REGION Network 3: Falha de comando
   RUNG wire#powerrail
      Contact( #TEMP0 )
      wire#w1
      S_Coil( #YFPP )
   END_RUNG
   RUNG wire#powerrail
      Contact( #TEMP1 )
   END_RUNG wire#w1
   RUNG wire#w1
      Coil( #AUX01 )
   END_RUNG
   // the same network as SCL:
   #_w1 := #TEMP0 OR #TEMP1;
   IF #_w1 THEN #YFPP := TRUE; END_IF;
   #AUX01 := #_w1;
END_REGION

REGION Network 4: Reset falha no acionamento
   RUNG wire#powerrail
      Contact( #CRF )
      I_Contact( #AUX01 )
      wire#w1
      R_Coil( #YFPP )
   END_RUNG
   RUNG wire#powerrail
      I_Contact( #DL )
   END_RUNG wire#w1
   // the same network as SCL:
   IF (#CRF AND NOT #AUX01) OR NOT #DL THEN #YFPP := FALSE; END_IF;
END_REGION

REGION Network 5: Falha
   RUNG wire#powerrail
      Contact( #DL )
      Contact( #MF1 )
      Contact( #MF2 )
      I_Contact( #YFPP )
      Not()
      Coil( #YF )
   END_RUNG
   // the same network as SCL:
   #YF := NOT (#DL AND #MF1 AND #MF2 AND NOT #YFPP);
END_REGION

REGION Network 6: Transição automático/manual
   RUNG wire#powerrail
      I_Contact( #CMA )
      P_Trig( #AUX02 )
      Contact( #MR )
      Contact( #ML )
      Coil( #AUX03 )
   END_RUNG
   // the same network as SCL:
   #_w1 := NOT #CMA AND NOT #AUX02;   // rising edge
   #AUX02 := NOT #CMA;
   #AUX03 := #_w1 AND #MR AND #ML;
END_REGION

REGION Network 7: Liga em manual
   RUNG wire#powerrail
      Contact( #CLM )
      wire#w1
      I_Contact( #CMA )
      I_Contact( #CDM )
      I_Contact( #YF )
      Contact( #HM )
      Contact( #MR )
      Coil( #AUX04 )
   END_RUNG
   RUNG wire#powerrail
      Contact( #AUX04 )
   END_RUNG wire#w1
   RUNG wire#powerrail
      Contact( #AUX03 )
   END_RUNG wire#w1
   // the same network as SCL:
   #AUX04 := (#CLM OR #AUX04 OR #AUX03) AND NOT #CMA AND NOT #CDM AND NOT #YF AND #HM AND #MR;
END_REGION

REGION Network 8: Liga em automático
   RUNG wire#powerrail
      Contact( #CMA )
      I_Contact( #YF )
      Contact( #HA )
      Contact( #MR )
      Coil( #AUX05 )
   END_RUNG
   // the same network as SCL:
   #AUX05 := #CMA AND NOT #YF AND #HA AND #MR;
END_REGION

REGION Network 9: Comando liga motor
   RUNG wire#powerrail
      Contact( #AUX05 )
      wire#w1
      Coil( #CL )
   END_RUNG
   RUNG wire#powerrail
      Contact( #AUX04 )
   END_RUNG wire#w1
   // the same network as SCL:
   #CL := #AUX05 OR #AUX04;
END_REGION

REGION Network 10
   RUNG wire#powerrail
      Contact( "AlwaysTRUE" )
      wire#w1
      Contact( #CL1S )
      Contact( #ML )
      P_Trig( #AUX06 )
      { S7_Templates := "SrcType := Int"; S7_GenerateENO := "TRUE" } Add(in1 := #SEG, in2 := 1, out => #SEG)
   END_RUNG
   RUNG wire#w1
      { S7_Templates := "SrcType := Int" } GE_Contact(in1 := #SEG, in2 := 60)
      P_Trig( #P60S )
      Coil( #AUX07 )
   END_RUNG
   // the same network as SCL:
   #_w1 := "AlwaysTRUE" AND #CL1S AND #ML;
   #_w2 := #_w1 AND NOT #AUX06;   // rising edge
   #AUX06 := #_w1;
   IF #_w2 THEN #SEG := #SEG + 1; END_IF;
   #_w3 := "AlwaysTRUE" AND (#SEG >= 60);
   #_w4 := #_w3 AND NOT #P60S;   // rising edge
   #P60S := #_w3;
   #AUX07 := #_w4;
END_REGION

REGION Network 11
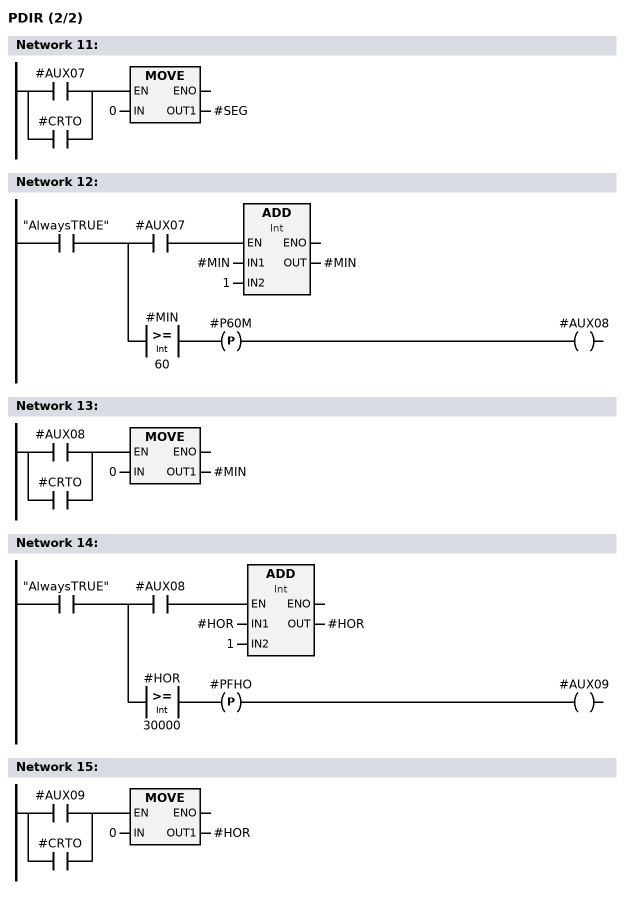
   RUNG wire#powerrail
      Contact( #AUX07 )
      wire#w1
      { S7_GenerateENO := "TRUE" } Move(in := 0, out1 => #SEG)
   END_RUNG
   RUNG wire#powerrail
      Contact( #CRTO )
   END_RUNG wire#w1
   // the same network as SCL:
   IF #AUX07 OR #CRTO THEN #SEG := 0; END_IF;
END_REGION

REGION Network 12
   RUNG wire#powerrail
      Contact( "AlwaysTRUE" )
      wire#w1
      Contact( #AUX07 )
      { S7_Templates := "SrcType := Int"; S7_GenerateENO := "TRUE" } Add(in1 := #MIN, in2 := 1, out => #MIN)
   END_RUNG
   RUNG wire#w1
      { S7_Templates := "SrcType := Int" } GE_Contact(in1 := #MIN, in2 := 60)
      P_Trig( #P60M )
      Coil( #AUX08 )
   END_RUNG
   // the same network as SCL:
   IF "AlwaysTRUE" AND #AUX07 THEN #MIN := #MIN + 1; END_IF;
   #_w1 := "AlwaysTRUE" AND (#MIN >= 60);
   #_w2 := #_w1 AND NOT #P60M;   // rising edge
   #P60M := #_w1;
   #AUX08 := #_w2;
END_REGION

REGION Network 13
   RUNG wire#powerrail
      Contact( #AUX08 )
      wire#w1
      { S7_GenerateENO := "TRUE" } Move(in := 0, out1 => #MIN)
   END_RUNG
   RUNG wire#powerrail
      Contact( #CRTO )
   END_RUNG wire#w1
   // the same network as SCL:
   IF #AUX08 OR #CRTO THEN #MIN := 0; END_IF;
END_REGION

REGION Network 14
   RUNG wire#powerrail
      Contact( "AlwaysTRUE" )
      wire#w1
      Contact( #AUX08 )
      { S7_Templates := "SrcType := Int"; S7_GenerateENO := "TRUE" } Add(in1 := #HOR, in2 := 1, out => #HOR)
   END_RUNG
   RUNG wire#w1
      { S7_Templates := "SrcType := Int" } GE_Contact(in1 := #HOR, in2 := 30000)
      P_Trig( #PFHO )
      Coil( #AUX09 )
   END_RUNG
   // the same network as SCL:
   IF "AlwaysTRUE" AND #AUX08 THEN #HOR := #HOR + 1; END_IF;
   #_w1 := "AlwaysTRUE" AND (#HOR >= 30000);
   #_w2 := #_w1 AND NOT #PFHO;   // rising edge
   #PFHO := #_w1;
   #AUX09 := #_w2;
END_REGION

REGION Network 15
   RUNG wire#powerrail
      Contact( #AUX09 )
      wire#w1
      { S7_GenerateENO := "TRUE" } Move(in := 0, out1 => #HOR)
   END_RUNG
   RUNG wire#powerrail
      Contact( #CRTO )
   END_RUNG wire#w1
   // the same network as SCL:
   IF #AUX09 OR #CRTO THEN #HOR := 0; END_IF;
END_REGION
END_FUNCTION_BLOCK

FUNCTION "ALARME" : Void   // FC2, SCL
{ S7_Optimized_Access := 'TRUE' }
VERSION : 0.1
BEGIN
   REGION "ALARMES IHM"
       // Statement section REGION
       "ALM0" := %DB300.DBW0;
       "ALM2" := %DB300.DBW2;
       "ALM4" := %DB300.DBW4;
       "ALM6" := %DB300.DBW6;
       "ALM8" := %DB300.DBW8;
       "ALM10" := %DB300.DBW10;
       "ALM12" := %DB300.DBW12;
       "ALM14" := %DB300.DBW14;
       "ALM16" := %DB300.DBW16;
   END_REGION
END_FUNCTION

FUNCTION "IO" : Void   // FC4, SCL
{ S7_Optimized_Access := 'TRUE' }
VERSION : 0.1
BEGIN
   REGION "Status e alarme elevatória principal 1"
       // Statement section REGION
       "Digitais"."MB-01-YFI" := "MB_01_DINV";
       "Digitais"."MB-01-YFB" := "MB_01_DMB";
       "Digitais"."MB-01-YFF" :="MB_01_FF";
       "Digitais"."MB-01-EMER" := NOT "MB_01_EMER";
       "Digitais"."MB-01-ML" :="MB_01_ML";
       "Digitais"."MB-01-YSH" :="MB_01_BL" OR "MB_01_SH";
       "Digitais"."MB-01-MM" :="MB_01_MMNT";
       "Digitais"."MB-01-MA" :="MB_01_MA";
       "Digitais"."MB-01-MN" :="MB_01_MN";
       "Digitais"."MB-01-HM" :="MB_01_HMNT";
       "Digitais"."MB-01-RST" :="MB_01_RST";
       "Digitais"."MB-01-INTRU" :="MB_01_INTRU";

       "MB_01_RR" :="COMANDOS"."MB-01-HS4";
       "MB_01_INTV" :="DIVERSOS"."MB-01-SP";
       "MB_01_INTVS" :="DIVERSOS"."MB-01-SP";


   END_REGION
   REGION "Status e alarme elevatória principal 2"
       // Statement section REGION
       "Digitais"."MB-02-YFI" := "MB_02_DINV";
       "Digitais"."MB-02-YFB" := "MB_02_DMB";
       "Digitais"."MB-02-YFF" := "MB_02_FF";
       "Digitais"."MB-02-EMER" := NOT "MB_02_EMER";
       "Digitais"."MB-02-ML" := "MB_02_ML";
       "Digitais"."MB-02-YSH" := "MB_02_BL" OR "MB_02_SH";
       "Digitais"."MB-02-MM" := "MB_02_MMNT";
       "Digitais"."MB-02-MA" := "MB_02_MA";
       "Digitais"."MB-02-MN" := "MB_02_MN";
       "Digitais"."MB-02-HM" := "MB_02_HMNT";
       "Digitais"."MB-02-RST" := "MB_02_RST";
       "Digitais"."MB-02-INTRU" := "MB_02_INTRU";

       "MB_02_RR" := "COMANDOS"."MB-02-HS4";
       "MB_02_INTV" := "DIVERSOS"."MB-02-SP";
       "MB_02_INTVS" := "DIVERSOS"."MB-02-SP";


   END_REGION
   REGION "Status e alarme elevatória principal 3"
       // Statement section REGION
       "Digitais"."MB-03-YFI" := "MB_03_DINV";
       "Digitais"."MB-03-YFB" := "MB_03_DMB";
       "Digitais"."MB-03-YFF" := "MB_03_FF";
       "Digitais"."MB-03-EMER" := NOT "MB_03_EMER";
       "Digitais"."MB-03-ML" := "MB_03_ML";
       "Digitais"."MB-03-YSH" := "MB_03_BL" OR "MB_03_SH";
       "Digitais"."MB-03-MM" := "MB_03_MMNT";
       "Digitais"."MB-03-MA" := "MB_03_MA";
       "Digitais"."MB-03-MN" := "MB_03_MN";
       "Digitais"."MB-03-HM" := "MB_03_HMNT";
       "Digitais"."MB-03-RST" := "MB_03_RST";
       "Digitais"."MB-03-INTRU" := "MB_03_INTRU";

       "MB_03_RR" := "COMANDOS"."MB-03-HS4";
       "MB_03_INTV" := "DIVERSOS"."MB-03-SP";
       "MB_03_INTVS" := "DIVERSOS"."MB-03-SP";


   END_REGION
   REGION "Status e alarme elevatória principal 4"
       // Statement section REGION
       "Digitais"."MB-04-YFI" := "MB_04_DINV";
       "Digitais"."MB-04-YFB" := "MB_04_DMB";
       "Digitais"."MB-04-YFF" := "MB_04_FF";
       "Digitais"."MB-04-EMER" := NOT "MB_04_EMER";
       "Digitais"."MB-04-ML" := "MB_04_ML";
       "Digitais"."MB-04-YSH" := "MB_04_BL" OR "MB_04_SH";
       "Digitais"."MB-04-MM" := "MB_04_MMNT";
       "Digitais"."MB-04-MA" := "MB_04_MA";
       "Digitais"."MB-04-MN" := "MB_04_MN";
       "Digitais"."MB-04-HM" := "MB_04_HMNT";
       "Digitais"."MB-04-RST" := "MB_04_RST";
       "Digitais"."MB-04-INTRU" := "MB_04_INTRU";

       "MB_04_RR" := "COMANDOS"."MB-04-HS4";
       "MB_04_INTV" := "DIVERSOS"."MB-04-SP";
       "MB_04_INTVS" := "DIVERSOS"."MB-04-SP";


   END_REGION

   REGION "Status e alarme PCM-E-CF-01-04"
       // Statement section REGION
       "Digitais".PCM_EEE_EMER := NOT "PCM_EEE_EMER";
       "Digitais".PCM_EEE_K27 := "PCM_EEE_K27";
       "Digitais".PCM_EEE_DISJ_LIG := "PCM_EEE_DJL";
       "Digitais".PCM_EEE_DISJ_DESLIG := "PCM_EEE_DJD";
       "Digitais".PCM_EEE_DISJ_YFAL := "PCM_EEE_DJYFAL";
       "Digitais".PCM_EEE_DISJ_FAL_GR := "PCM_EEE_DJFG";
       "Digitais".PCM_EEE_TR01_KA3 := "PCM_EEE_TR01_KA3";
       "Digitais".PCM_EEE_TR01_KA4 := "PCM_EEE_TR01_KA4";
       "Digitais".PCM_EEE_TR01_KA5 := "PCM_EEE_TR01_KA5";
       "Digitais".PCM_EEE_INTRU := "PCM_EEE_INTRU";
   END_REGION

   REGION "Status e alarme QGBT-AUX-01"
       // Statement section REGION
       "Digitais".QGBT_EMER := NOT "QGBT_EMER";
       "Digitais".QGBT_K27 := "QGBT_K27";
       "Digitais".QGBT_DJL := "QGBT_DISJ_LIG";
       "Digitais".QGBT_DJD := "QGBT_DISJ_DESLIG";
       "Digitais".QGBT_DJYFAL := "QGBT_DISJ_YFAL";
       "Digitais".QGBT_INTRU := "QGBT_INTRU";
   END_REGION

   REGION "CHAVE DE NIVEL LS-001"
       // Statement section REGION
       // 
       "DIVERSOS".TMR[5].TON(IN := "LSL_001",
                             PT := T#5S);
       "DIVERSOS".TMR[6].TON(IN := "LSH_001",
                             PT := T#5S);
       "Digitais".LSL_001 := "DIVERSOS".TMR[5].Q;
       "Digitais".LSH_001 := "DIVERSOS".TMR[6].Q;
   END_REGION

   REGION "CHAVE DE NIVEL LS-002"
       // Statement section REGION
       "DIVERSOS".TMR[7].TON(IN := "LSL_002",
                             PT := T#5S);
       "DIVERSOS".TMR[8].TON(IN := "LSH_002",
                             PT := T#5S);
       "Digitais".LSL_002 := "DIVERSOS".TMR[7].Q;
       "Digitais".LSH_002 := "DIVERSOS".TMR[8].Q;
   END_REGION

   REGION "Status e alarme PCE-EEE"
       // Statement section REGION
       "Digitais".PCE_EEE_INTRU := "PCE_EEE_INTRU";
       "Digitais".PCE_EEE_UPS_ALM := "PCE_EEE_UPS_ALM";
       "Digitais".PCE_EEE_UPS_FE := "PCE_EEE_UPS_FE";
       "Digitais".PCE_EEE_UPS_CHAR := "PCE_EEE_UPS_CHAR";






   END_REGION
END_FUNCTION

FUNCTION "MB-01" : Void   // FC7, SCL
{ S7_Optimized_Access := 'TRUE' }
VERSION : 0.1
   VAR_TEMP
      IM : Bool;   // Intertravamento manual = 0
      IA : Bool;   // Intertravamento automáticol = 0
      HABM : Bool;   // Habilita funcionamento manual = 1
      HABA : Bool;   // Habilita funcionamento automático = 1
      CLM : Bool;   // Comando liga motor
      PROT : Bool;   // Proteção do motor acionada
   END_VAR
BEGIN
   REGION Intertravamento maual/automático
       // Statement section REGION
       IF (NOT "Digitais".QGBT_EMER AND NOT "Digitais".PCM_EEE_EMER AND NOT "Digitais"."MB-01-EMER") = 1 THEN
           // Statement section IF
           #IA := 1;
           #IM := 1;
       ELSE
           #IA := 0;
           #IM := 0;
       END_IF;

   END_REGION

   REGION Habilita funcionamento automático
       // Statement section REGION
       IF (#IA AND "DIVERSOS"."MB-01-SP") = 1 THEN
           // Statement section IF
           #HABA := 1;
       ELSE
           #HABA := 0;
       END_IF;

   END_REGION

   REGION Habilita funcionamento manual
       // Statement section REGION
       IF #IM THEN
           // Statement section IF
           #HABM := 1;
       ELSE
           #HABM := 0;
       END_IF;
   END_REGION

   REGION Bloco de acionamento DO motor
       // Statement section REGION
       "PDIR_DB_MB-01"(ML:="Digitais"."MB-01-YSH",
                       MR:="Digitais"."MB-01-YR",
                       DL:=NOT "Digitais"."MB-01-YFI" AND NOT "Digitais"."MB-01-YFB" AND NOT "Digitais"."MB-01-YFF",
                       MF1:="AlwaysTRUE",
                       MF2:="AlwaysTRUE",
                       HM:=#HABM,
                       HA:=#HABA,
                       CMA:="COMANDOS"."MB-01-HS1",
                       CLM:="COMANDOS"."MB-01-HS2",
                       CDM:="COMANDOS"."MB-01-HS3",
                       CRF:="COMANDOS"."MB-01-HS4" OR "Digitais"."MB-01-RST",
                       CRTO:="COMANDOS"."MB-01-HS5",
                       CL1S:="Clock_1Hz",
                       YFPP=>"Digitais"."MB-01-YFA",
                       YF=>"Digitais"."MB-01-YF",
                       CL=>"MB_01_SH",
                       SEG:="Totalizadores"."MB-01-SO",
                       MIN:="Totalizadores"."MB-01-MO",
                       HOR:="Totalizadores"."MB-01-HO");

                    END_REGION

   REGION Reset dos comandos de pulso
       // Statement section REGION
       IF "COMANDOS"."MB-01-HS2" THEN
           // Statement section IF
           "COMANDOS"."MB-01-HS2" := 0;
       END_IF;
       IF "COMANDOS"."MB-01-HS3" THEN
           // Statement section IF
           "COMANDOS"."MB-01-HS3" := 0;
       END_IF;
       IF "COMANDOS"."MB-01-HS4" THEN
           // Statement section IF
           "COMANDOS"."MB-01-HS4" := 0;
       END_IF;
       IF "COMANDOS"."MB-01-HS5" THEN
           // Statement section IF
           "COMANDOS"."MB-01-HS5" := 0;
       END_IF;
   END_REGION

   REGION Elevatoria principal modo automatico
       IF ("Digitais"."MB-01-MA") = 1 THEN
           "Digitais"."MB-01-YR" := 1;
       ELSE
           "Digitais"."MB-01-YR" := 0;
       END_IF;

   END_REGION

   REGION Proteção hidraulica MB-01
       // Statement section REGION
       IF ("VARIAVEIS".LIT_001 <= "SETPOINTS".SP_NVL_MIN) OR "Digitais".LSL_002 OR "Digitais"."LIT_001-YLL" THEN
           // Statement section IF
           "MB_01_PH" := 1;
       ELSE
           "MB_01_PH" := 0;
       END_IF;

   END_REGION
END_FUNCTION

FUNCTION "MB-02" : Void   // FC8, SCL
{ S7_Optimized_Access := 'TRUE' }
VERSION : 0.1
   VAR_TEMP
      IM : Bool;   // Intertravamento manual = 0
      IA : Bool;   // Intertravamento automáticol = 0
      HABM : Bool;   // Habilita funcionamento manual = 1
      HABA : Bool;   // Habilita funcionamento automático = 1
      CLM : Bool;   // Comando liga motor
      PROT : Bool;   // Proteção do motor acionada
   END_VAR
BEGIN
   REGION Intertravamento maual/automático
       // Statement section REGION
       IF (NOT "Digitais".QGBT_EMER AND NOT "Digitais".PCM_EEE_EMER AND NOT "Digitais"."MB-02-EMER") = 1 THEN
           // Statement section IF
           #IA := 1;
           #IM := 1;
       ELSE
           #IA := 0;
           #IM := 0;
       END_IF;

   END_REGION

   REGION Habilita funcionamento automático
       // Statement section REGION
       IF (#IA AND "DIVERSOS"."MB-02-SP") = 1 THEN
           // Statement section IF
           #HABA := 1;
       ELSE
           #HABA := 0;
       END_IF;

   END_REGION

   REGION Habilita funcionamento manual
       // Statement section REGION
       IF #IM THEN
           // Statement section IF
           #HABM := 1;
       ELSE
           #HABM := 0;
       END_IF;
   END_REGION

   REGION Bloco de acionamento DO motor
       // Statement section REGION
       "PDIR_DB_MB-02"(ML:="Digitais"."MB-02-YSH",
                       MR:="Digitais"."MB-02-MA",
                       DL:=NOT "Digitais"."MB-02-YFI" AND NOT "Digitais"."MB-02-YFB" AND NOT "Digitais"."MB-02-YFF",
                       MF1:="AlwaysTRUE",
                       MF2:="AlwaysTRUE",
                       HM:=#HABM,
                       HA:=#HABA,
                       CMA:="COMANDOS"."MB-02-HS1",
                       CLM:="COMANDOS"."MB-02-HS2",
                       CDM:="COMANDOS"."MB-02-HS3",
                       CRF:="COMANDOS"."MB-02-HS4" OR "Digitais"."MB-02-RST",
                       CRTO:="COMANDOS"."MB-02-HS5",
                       CL1S:="Clock_1Hz",
                       YFPP=>"Digitais"."MB-02-YFA",
                       YF=>"Digitais"."MB-02-YF",
                       CL=>"MB_02_SH",
                       SEG:="Totalizadores"."MB-02-SO",
                       MIN:="Totalizadores"."MB-02-MO",
                       HOR:="Totalizadores"."MB-02-HO");

                    END_REGION

   REGION Reset dos comandos de pulso
       // Statement section REGION
       IF "COMANDOS"."MB-02-HS2" THEN
           // Statement section IF
           "COMANDOS"."MB-02-HS2" := 0;
       END_IF;
       IF "COMANDOS"."MB-02-HS3" THEN
           // Statement section IF
           "COMANDOS"."MB-02-HS3" := 0;
       END_IF;
       IF "COMANDOS"."MB-02-HS4" THEN
           // Statement section IF
           "COMANDOS"."MB-02-HS4" := 0;
       END_IF;
       IF "COMANDOS"."MB-02-HS5" THEN
           // Statement section IF
           "COMANDOS"."MB-02-HS5" := 0;
       END_IF;
   END_REGION

   REGION Elevatoria principal modo automatico
       "Digitais"."MB-02-YR" := "Digitais"."MB-02-MA";
   END_REGION

   REGION Proteção hidraulica MB-02
       // Statement section REGION
       IF ("VARIAVEIS".LIT_001 <= "SETPOINTS".SP_NVL_MIN) OR "Digitais".LSL_002 OR "Digitais"."LIT_001-YLL" THEN
           // Statement section IF
           "MB_02_PH" := 1;
       ELSE
           "MB_02_PH" := 0;
       END_IF;

   END_REGION
END_FUNCTION

FUNCTION "MB-03" : Void   // FC9, SCL
{ S7_Optimized_Access := 'TRUE' }
VERSION : 0.1
   VAR_TEMP
      IM : Bool;   // Intertravamento manual = 0
      IA : Bool;   // Intertravamento automáticol = 0
      HABM : Bool;   // Habilita funcionamento manual = 1
      HABA : Bool;   // Habilita funcionamento automático = 1
      CLM : Bool;   // Comando liga motor
      PROT : Bool;   // Proteção do motor acionada
   END_VAR
BEGIN
   REGION Intertravamento maual/automático
       // Statement section REGION
       IF (NOT "Digitais".QGBT_EMER AND NOT "Digitais".PCM_EEE_EMER AND NOT "Digitais"."MB-03-EMER") = 1 THEN
           // Statement section IF
           #IA := 1;
           #IM := 1;
       ELSE
           #IA := 0;
           #IM := 0;
       END_IF;

   END_REGION

   REGION Habilita funcionamento automático
       // Statement section REGION
       IF (#IA AND "DIVERSOS"."MB-03-SP") = 1 THEN
           // Statement section IF
           #HABA := 1;
       ELSE
           #HABA := 0;
       END_IF;

   END_REGION

   REGION Habilita funcionamento manual
       // Statement section REGION
       IF #IM THEN
           // Statement section IF
           #HABM := 1;
       ELSE
           #HABM := 0;
       END_IF;
   END_REGION

   REGION Bloco de acionamento DO motor
       // Statement section REGION
       "PDIR_DB_MB-03"(ML:="Digitais"."MB-03-YSH",
                       MR:="Digitais"."MB-03-MA",
                       DL:=NOT "Digitais"."MB-03-YFI" AND NOT "Digitais"."MB-03-YFB" AND NOT "Digitais"."MB-03-YFF",
                       MF1:="AlwaysTRUE",
                       MF2:="AlwaysTRUE",
                       HM:=#HABM,
                       HA:=#HABA,
                       CMA:="COMANDOS"."MB-03-HS1",
                       CLM:="COMANDOS"."MB-03-HS2",
                       CDM:="COMANDOS"."MB-03-HS3",
                       CRF:="COMANDOS"."MB-03-HS4" OR "Digitais"."MB-03-RST",
                       CRTO:="COMANDOS"."MB-03-HS5",
                       CL1S:="Clock_1Hz",
                       YFPP=>"Digitais"."MB-03-YFA",
                       YF=>"Digitais"."MB-03-YF",
                       CL=>"MB_03_SH",
                       SEG:="Totalizadores"."MB-03-SO",
                       MIN:="Totalizadores"."MB-03-MO",
                       HOR:="Totalizadores"."MB-03-HO");

                    END_REGION

   REGION Reset dos comandos de pulso
       // Statement section REGION
       IF "COMANDOS"."MB-03-HS2" THEN
           // Statement section IF
           "COMANDOS"."MB-03-HS2" := 0;
       END_IF;
       IF "COMANDOS"."MB-03-HS3" THEN
           // Statement section IF
           "COMANDOS"."MB-03-HS3" := 0;
       END_IF;
       IF "COMANDOS"."MB-03-HS4" THEN
           // Statement section IF
           "COMANDOS"."MB-03-HS4" := 0;
       END_IF;
       IF "COMANDOS"."MB-03-HS5" THEN
           // Statement section IF
           "COMANDOS"."MB-03-HS5" := 0;
       END_IF;
   END_REGION

   REGION Elevatoria principal modo automatico
       "Digitais"."MB-03-YR" := "Digitais"."MB-03-MA";
   END_REGION

   REGION Proteção hidraulica MB-03
       // Statement section REGION
       IF ("VARIAVEIS".LIT_001 <= "SETPOINTS".SP_NVL_MIN) OR "Digitais".LSL_002 OR "Digitais"."LIT_001-YLL" THEN
           // Statement section IF
           "MB_03_PH" := 1;
       ELSE
           "MB_03_PH" := 0;
       END_IF;

   END_REGION
END_FUNCTION

FUNCTION "MB-04" : Void   // FC10, SCL
{ S7_Optimized_Access := 'TRUE' }
VERSION : 0.1
   VAR_TEMP
      IM : Bool;   // Intertravamento manual = 0
      IA : Bool;   // Intertravamento automáticol = 0
      HABM : Bool;   // Habilita funcionamento manual = 1
      HABA : Bool;   // Habilita funcionamento automático = 1
      CLM : Bool;   // Comando liga motor
      PROT : Bool;   // Proteção do motor acionada
   END_VAR
BEGIN
   REGION Intertravamento maual/automático
       // Statement section REGION
       IF (NOT "Digitais".QGBT_EMER AND NOT "Digitais".PCM_EEE_EMER AND NOT "Digitais"."MB-04-EMER") = 1 THEN
           // Statement section IF
           #IA := 1;
           #IM := 1;
       ELSE
           #IA := 0;
           #IM := 0;
       END_IF;

   END_REGION

   REGION Habilita funcionamento automático
       // Statement section REGION
       IF (#IA AND "DIVERSOS"."MB-04-SP") = 1 THEN
           // Statement section IF
           #HABA := 1;
       ELSE
           #HABA := 0;
       END_IF;

   END_REGION

   REGION Habilita funcionamento manual
       // Statement section REGION
       IF #IM THEN
           // Statement section IF
           #HABM := 1;
       ELSE
           #HABM := 0;
       END_IF;
   END_REGION

   REGION Bloco de acionamento DO motor
       // Statement section REGION
       "PDIR_DB_MB-04"(ML:="Digitais"."MB-04-YSH",
                       MR:="Digitais"."MB-04-MA",
                       DL:=NOT "Digitais"."MB-04-YFI" AND NOT "Digitais"."MB-04-YFB" AND NOT "Digitais"."MB-04-YFF",
                       MF1:="AlwaysTRUE",
                       MF2:="AlwaysTRUE",
                       HM:=#HABM,
                       HA:=#HABA,
                       CMA:="COMANDOS"."MB-04-HS1",
                       CLM:="COMANDOS"."MB-04-HS2",
                       CDM:="COMANDOS"."MB-04-HS3",
                       CRF:="COMANDOS"."MB-04-HS4" OR "Digitais"."MB-04-RST",
                       CRTO:="COMANDOS"."MB-04-HS5",
                       CL1S:="Clock_1Hz",
                       YFPP=>"Digitais"."MB-04-YFA",
                       YF=>"Digitais"."MB-04-YF",
                       CL=>"MB_04_SH",
                       SEG:="Totalizadores"."MB-04-SO",
                       MIN:="Totalizadores"."MB-04-MO",
                       HOR:="Totalizadores"."MB-04-HO");

                    END_REGION

   REGION Reset dos comandos de pulso
       // Statement section REGION
       IF "COMANDOS"."MB-04-HS2" THEN
           // Statement section IF
           "COMANDOS"."MB-04-HS2" := 0;
       END_IF;
       IF "COMANDOS"."MB-04-HS3" THEN
           // Statement section IF
           "COMANDOS"."MB-04-HS3" := 0;
       END_IF;
       IF "COMANDOS"."MB-04-HS4" THEN
           // Statement section IF
           "COMANDOS"."MB-04-HS4" := 0;
       END_IF;
       IF "COMANDOS"."MB-04-HS5" THEN
           // Statement section IF
           "COMANDOS"."MB-04-HS5" := 0;
       END_IF;
   END_REGION

   REGION Elevatoria principal modo automatico
       "Digitais"."MB-04-YR" := "Digitais"."MB-04-MA";
   END_REGION

   REGION Proteção hidraulica MB-04
       // Statement section REGION
       IF ("VARIAVEIS".LIT_001 <= "SETPOINTS".SP_NVL_MIN) OR "Digitais".LSL_002 OR "Digitais"."LIT_001-YLL" THEN
           // Statement section IF
           "MB_04_PH" := 1;
       ELSE
           "MB_04_PH" := 0;
       END_IF;

   END_REGION
END_FUNCTION

ORGANIZATION_BLOCK "Main"   // OB1, LAD, ProgramCycle
TITLE = "Main Program Sweep (Cycle)"
{ S7_Optimized_Access := 'TRUE' }
VERSION : 0.1
   VAR_INPUT
      Initial_Call : Bool;   // Initial call of this OB
      Remanence : Bool;   // =True, if remanent data are available
   END_VAR
BEGIN

REGION Network 1: PULSO 1 SEGUNDO
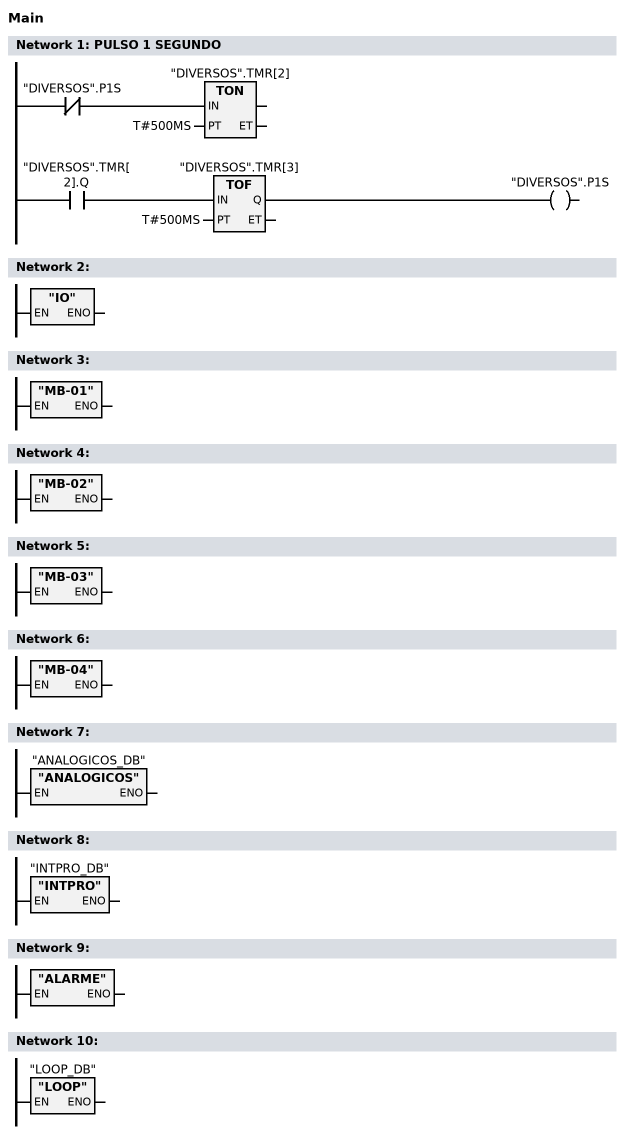
   "DIVERSOS".TMR[2].TON(IN := NOT "DIVERSOS".P1S, PT := T#500MS);
   "DIVERSOS".TMR[3].TOF(IN := "DIVERSOS".TMR[2].Q, PT := T#500MS);
   "DIVERSOS".P1S := "DIVERSOS".TMR[3].Q;
END_REGION

REGION Network 2
   RUNG wire#powerrail
      "IO"()
   END_RUNG
   // the same network as SCL:
   "IO"();
END_REGION

REGION Network 3
   RUNG wire#powerrail
      "MB-01"()
   END_RUNG
   // the same network as SCL:
   "MB-01"();
END_REGION

REGION Network 4
   RUNG wire#powerrail
      "MB-02"()
   END_RUNG
   // the same network as SCL:
   "MB-02"();
END_REGION

REGION Network 5
   RUNG wire#powerrail
      "MB-03"()
   END_RUNG
   // the same network as SCL:
   "MB-03"();
END_REGION

REGION Network 6
   RUNG wire#powerrail
      "MB-04"()
   END_RUNG
   // the same network as SCL:
   "MB-04"();
END_REGION

REGION Network 7
   RUNG wire#powerrail
      "ANALOGICOS_DB"()
   END_RUNG
   // the same network as SCL:
   "ANALOGICOS_DB"();   // "ANALOGICOS"
END_REGION

REGION Network 8
   RUNG wire#powerrail
      "INTPRO_DB"()
   END_RUNG
   // the same network as SCL:
   "INTPRO_DB"();   // "INTPRO"
END_REGION

REGION Network 9
   RUNG wire#powerrail
      "ALARME"()
   END_RUNG
   // the same network as SCL:
   "ALARME"();
END_REGION

REGION Network 10
   RUNG wire#powerrail
      "LOOP_DB"()
   END_RUNG
   // the same network as SCL:
   "LOOP_DB"();   // "LOOP"
END_REGION
END_ORGANIZATION_BLOCK

ORGANIZATION_BLOCK "Cyclic interrupt"   // OB30, SCL, CyclicInterrupt
{ S7_Optimized_Access := 'TRUE' }
VERSION : 0.1
   VAR_INPUT
      Initial_Call : Bool;   // Initial call of this OB
      Event_Count : Int;   // Events discarded
   END_VAR
   VAR_TEMP
      OB35_EV_CLASS : Byte;
      OB35_STRT_INF : Byte;
      OB35_PRIORITY : Byte;
      OB35_OB_NUMBR : Byte;
      OB35_RESERVED_1 : Byte;
      OB35_RESERVED_2 : Byte;
      OB35_PHASE_OFFSET : Word;
      OB35_RESERVED_3 : Int;
      OB35_EXC_FREQ : Int;
      OB35_DATE_TIME : Date_And_Time;
      "SPM-EEEB" : Real;   // Setpoint manual PID tanque de aeração 1
      EEEB_IT : Time;   // Ajuste integral do PID
      EEEB_DT : Time;   // Ajuste derivativo do PID
      EEEB_AUX : Real;   // Setpoint manual PID - auxiliar
      EEEB_P : Real;   // Setpoint manual PID - auxiliar
      AUX1 : Real;
   END_VAR
BEGIN
   REGION CONVERSÃO DOS SETPOINTS PARA TEMPO PID EEEB
       // Statement section REGION
       #EEEB_IT := ROUND(("PID"."PID-EEEB-I" * 1000.0));

       #EEEB_DT := ROUND(("PID"."PID-EEEB-D" * 1000.0));

       #EEEB_P := "PID"."PID-EEEB-P" * -1;
   END_REGION
   REGION "PID" TANQUE
       // Statement section REGION
       "PID-EEEB"(MAN_ON:="COMANDOS"."PID-EEEB-HM",
                  P_SEL:="COMANDOS"."PID-EEEB-HP",
                  I_SEL:="COMANDOS"."PID-EEEB-HI",
                  D_SEL:="COMANDOS"."PID-EEEB-HD",
                  CYCLE:=T#30S,
                  SP_INT:="SETPOINTS"."LIT_001-SPC",
                  PV_IN:="VARIAVEIS"."LIT_001-P",
                  MAN:="PID"."PID-EEEB-SPM",
                  GAIN:=#EEEB_P,
                  TI:=#EEEB_IT,
                  TD:=#EEEB_DT,
                  DEADB_W:="PID"."PID-EEEB-DB",
                  LMN_HLM:="PID"."PID-EEEB-MAX",
                  LMN_LLM:="PID"."PID-EEEB-MIN",
                  PV_FAC := 1.0,
                  LMN=>"PID"."VA-PID-EEEB");


   END_REGION
   REGION Valor Relativo
       // Statement section REGION
       "PID"."PID-EEEB-VR" := "SETPOINTS"."LIT_001-SPC" / "VARIAVEIS"."LIT_001-P";
   END_REGION
   REGION Calculo para encontrar fator de multiplicação 
       // Statement section REGION
       "PID".AUX_CALC[5] := 27648.0 / "PID"."PID-EEEB-MAX";
   END_REGION
   REGION Movimenta saida PID para entrada analógica inversor
       //MOVIMENTA PARA SAIDA ANALOGICA MB-01
       IF "Digitais"."MB-01-YSH" THEN
           // Statement section IF
           "MB_01_VEL" := REAL_TO_INT("PID".AUX_CALC[1]);
           IF "COMANDOS"."MB-01-HS1" THEN
               // Statement section IF
               "PID".AUX_CALC[1] := "PID"."VA-PID-EEEB" * "PID".AUX_CALC[5];
           ELSE
               "PID".AUX_CALC[1] := "SETPOINTS"."MB-01-SP" * "PID".AUX_CALC[5];
           END_IF;
       END_IF;

       //MOVIMENTA PARA SAIDA ANALOGICA MB-02
       IF "Digitais"."MB-02-YSH" THEN
           // Statement section IF
           "MB_02_VEL" := REAL_TO_INT("PID".AUX_CALC[2]);
           IF "COMANDOS"."MB-02-HS1" THEN
               // Statement section IF
               "PID".AUX_CALC[2] := "PID"."VA-PID-EEEB" * "PID".AUX_CALC[5];
           ELSE
               "PID".AUX_CALC[2] := "SETPOINTS"."MB-02-SP" * "PID".AUX_CALC[5];
           END_IF;
       END_IF;

       //MOVIMENTA PARA SAIDA ANALOGICA MB-03
       IF "Digitais"."MB-03-YSH" THEN
           "MB_03_VEL" := REAL_TO_INT("PID".AUX_CALC[3]);
           IF "COMANDOS"."MB-03-HS1" THEN
               "PID".AUX_CALC[3] := "PID"."VA-PID-EEEB" * "PID".AUX_CALC[5];
           ELSE
               "PID".AUX_CALC[3] := "SETPOINTS"."MB-03-SP" * "PID".AUX_CALC[5];
           END_IF;
       END_IF;

       //MOVIMENTA PARA SAIDA ANALOGICA MB-04
       IF "Digitais"."MB-04-YSH" THEN
           // Statement section IF
           "MB_04_VEL" := REAL_TO_INT("PID".AUX_CALC[4]);
           IF "COMANDOS"."MB-03-HS1" THEN
               // Statement section IF
               "PID".AUX_CALC[4] := "PID"."VA-PID-EEEB" * "PID".AUX_CALC[5];
           ELSE
               "PID".AUX_CALC[4] := "SETPOINTS"."MB-04-SP" * "PID".AUX_CALC[5];
           END_IF;
       END_IF;
   END_REGION
END_ORGANIZATION_BLOCK

(* ===== HMI "HMI_RT_1" =====
system functions are stored by id; their names below are inferred from use
connection "HMI_Connection_1": ETHERNET, SMART_S7_1500_OMS

HMI tags "Default tag table"
   "Digitais_MB-01-YSH" : Bool = PLC Digitais.MB-01-YSH AT %DB300.DBX0.0, 1 s
   "pause" : Bool = PLC pause AT %M2.1, 1 s
   "DIVERSOS_Looping" : Int = PLC DIVERSOS.Looping, 1 s
   "Tag_ScreenNumber" : Int, internal

HMI tags "ALARMES"
   "ALM0" : Word = PLC ALM0 AT %MW100, 1 s
   "ALM2" : Word = PLC ALM2 AT %MW102, 1 s
   "ALM4" : Word = PLC ALM4 AT %MW104, 1 s
   "ALM6" : Word = PLC ALM6 AT %MW106, 1 s
   "ALM8" : Word = PLC ALM8 AT %MW108, 1 s
   "ALM10" : Word = PLC ALM10 AT %MW110, 1 s
   "ALM12" : Word = PLC ALM12 AT %MW112, 1 s
   "ALM14" : Word = PLC ALM14 AT %MW114, 1 s
   "ALM16" : Word = PLC ALM16 AT %MW116, 1 s

HMI tags "PID"
   "PID_PID-EEEB-D" : Real = PLC PID.PID-EEEB-D AT %DB307.DBD0, 1 s
   "PID_PID-EEEB-P" : Real = PLC PID.PID-EEEB-P AT %DB307.DBD4, 1 s
   "PID_PID-EEEB-I" : Real = PLC PID.PID-EEEB-I AT %DB307.DBD8, 1 s
   "PID_PID-EEEB-MIN" : Real = PLC PID.PID-EEEB-MIN AT %DB307.DBD12, 1 s
   "PID_PID-EEEB-MAX" : Real = PLC PID.PID-EEEB-MAX AT %DB307.DBD16, 1 s
   "PID_PID-EEEB-DB" : Real = PLC PID.PID-EEEB-DB AT %DB307.DBD20, 1 s
   "PID_PID-EEEB-SPM" : Real = PLC PID.PID-EEEB-SPM AT %DB307.DBD24, 1 s
   "PID_VA-PID-EEEB" : Real = PLC PID.VA-PID-EEEB AT %DB307.DBD28, 1 s
   "PID_PID-EEEB-VR" : Real = PLC PID.PID-EEEB-VR AT %DB307.DBD32, 1 s

HMI tags "Comandos"
   "COMANDOS_MB-01-HS9" : Bool = PLC COMANDOS.MB-01-HS9 AT %DB303.DBX0.0, 1 s
   "COMANDOS_MB-01-HS10" : Bool = PLC COMANDOS.MB-01-HS10 AT %DB303.DBX0.1, 1 s
   "COMANDOS_MB-01-HS11" : Bool = PLC COMANDOS.MB-01-HS11 AT %DB303.DBX0.2, 1 s
   "COMANDOS_MB-01-HS12" : Bool = PLC COMANDOS.MB-01-HS12 AT %DB303.DBX0.3, 1 s
   "COMANDOS_MB-01-HS13" : Bool = PLC COMANDOS.MB-01-HS13 AT %DB303.DBX0.4, 1 s
   "COMANDOS_MB-01-HS14" : Bool = PLC COMANDOS.MB-01-HS14 AT %DB303.DBX0.5, 1 s
   "COMANDOS_MB-01-HS15" : Bool = PLC COMANDOS.MB-01-HS15 AT %DB303.DBX0.6, 1 s
   "COMANDOS_MB-01-HS16" : Bool = PLC COMANDOS.MB-01-HS16 AT %DB303.DBX0.7, 1 s
   "COMANDOS_MB-01-HS1" : Bool = PLC COMANDOS.MB-01-HS1 AT %DB303.DBX1.0, 1 s
   "COMANDOS_MB-01-HS2" : Bool = PLC COMANDOS.MB-01-HS2 AT %DB303.DBX1.1, 1 s
   "COMANDOS_MB-01-HS3" : Bool = PLC COMANDOS.MB-01-HS3 AT %DB303.DBX1.2, 1 s
   "COMANDOS_MB-01-HS4" : Bool = PLC COMANDOS.MB-01-HS4 AT %DB303.DBX1.3, 1 s
   "COMANDOS_MB-01-HS5" : Bool = PLC COMANDOS.MB-01-HS5 AT %DB303.DBX1.4, 1 s
   "COMANDOS_MB-01-HS6" : Bool = PLC COMANDOS.MB-01-HS6 AT %DB303.DBX1.5, 1 s
   "COMANDOS_MB-01-HS7" : Bool = PLC COMANDOS.MB-01-HS7 AT %DB303.DBX1.6, 1 s
   "COMANDOS_MB-01-HS8" : Bool = PLC COMANDOS.MB-01-HS8 AT %DB303.DBX1.7, 1 s
   "COMANDOS_MB-02-HS9" : Bool = PLC COMANDOS.MB-02-HS9 AT %DB303.DBX2.0, 1 s
   "COMANDOS_MB-02-HS10" : Bool = PLC COMANDOS.MB-02-HS10 AT %DB303.DBX2.1, 1 s
   "COMANDOS_MB-02-HS11" : Bool = PLC COMANDOS.MB-02-HS11 AT %DB303.DBX2.2, 1 s
   "COMANDOS_MB-02-HS12" : Bool = PLC COMANDOS.MB-02-HS12 AT %DB303.DBX2.3, 1 s
   "COMANDOS_MB-02-HS13" : Bool = PLC COMANDOS.MB-02-HS13 AT %DB303.DBX2.4, 1 s
   "COMANDOS_MB-02-HS14" : Bool = PLC COMANDOS.MB-02-HS14 AT %DB303.DBX2.5, 1 s
   "COMANDOS_MB-02-HS15" : Bool = PLC COMANDOS.MB-02-HS15 AT %DB303.DBX2.6, 1 s
   "COMANDOS_MB-02-HS16" : Bool = PLC COMANDOS.MB-02-HS16 AT %DB303.DBX2.7, 1 s
   "COMANDOS_MB-02-HS1" : Bool = PLC COMANDOS.MB-02-HS1 AT %DB303.DBX3.0, 1 s
   "COMANDOS_MB-02-HS2" : Bool = PLC COMANDOS.MB-02-HS2 AT %DB303.DBX3.1, 1 s
   "COMANDOS_MB-02-HS3" : Bool = PLC COMANDOS.MB-02-HS3 AT %DB303.DBX3.2, 1 s
   "COMANDOS_MB-02-HS4" : Bool = PLC COMANDOS.MB-02-HS4 AT %DB303.DBX3.3, 1 s
   "COMANDOS_MB-02-HS5" : Bool = PLC COMANDOS.MB-02-HS5 AT %DB303.DBX3.4, 1 s
   "COMANDOS_MB-02-HS6" : Bool = PLC COMANDOS.MB-02-HS6 AT %DB303.DBX3.5, 1 s
   "COMANDOS_MB-02-HS7" : Bool = PLC COMANDOS.MB-02-HS7 AT %DB303.DBX3.6, 1 s
   "COMANDOS_MB-02-HS8" : Bool = PLC COMANDOS.MB-02-HS8 AT %DB303.DBX3.7, 1 s
   "COMANDOS_MB-03-HS9" : Bool = PLC COMANDOS.MB-03-HS9 AT %DB303.DBX4.0, 1 s
   "COMANDOS_MB-03-HS10" : Bool = PLC COMANDOS.MB-03-HS10 AT %DB303.DBX4.1, 1 s
   "COMANDOS_MB-03-HS11" : Bool = PLC COMANDOS.MB-03-HS11 AT %DB303.DBX4.2, 1 s
   "COMANDOS_MB-03-HS12" : Bool = PLC COMANDOS.MB-03-HS12 AT %DB303.DBX4.3, 1 s
   "COMANDOS_MB-03-HS13" : Bool = PLC COMANDOS.MB-03-HS13 AT %DB303.DBX4.4, 1 s
   "COMANDOS_MB-03-HS14" : Bool = PLC COMANDOS.MB-03-HS14 AT %DB303.DBX4.5, 1 s
   "COMANDOS_MB-03-HS15" : Bool = PLC COMANDOS.MB-03-HS15 AT %DB303.DBX4.6, 1 s
   "COMANDOS_MB-03-HS16" : Bool = PLC COMANDOS.MB-03-HS16 AT %DB303.DBX4.7, 1 s
   "COMANDOS_MB-03-HS1" : Bool = PLC COMANDOS.MB-03-HS1 AT %DB303.DBX5.0, 1 s
   "COMANDOS_MB-03-HS2" : Bool = PLC COMANDOS.MB-03-HS2 AT %DB303.DBX5.1, 1 s
   "COMANDOS_MB-03-HS3" : Bool = PLC COMANDOS.MB-03-HS3 AT %DB303.DBX5.2, 1 s
   "COMANDOS_MB-03-HS4" : Bool = PLC COMANDOS.MB-03-HS4 AT %DB303.DBX5.3, 1 s
   "COMANDOS_MB-03-HS5" : Bool = PLC COMANDOS.MB-03-HS5 AT %DB303.DBX5.4, 1 s
   "COMANDOS_MB-03-HS6" : Bool = PLC COMANDOS.MB-03-HS6 AT %DB303.DBX5.5, 1 s
   "COMANDOS_MB-03-HS7" : Bool = PLC COMANDOS.MB-03-HS7 AT %DB303.DBX5.6, 1 s
   "COMANDOS_MB-03-HS8" : Bool = PLC COMANDOS.MB-03-HS8 AT %DB303.DBX5.7, 1 s
   "COMANDOS_MB-04-HS9" : Bool = PLC COMANDOS.MB-04-HS9 AT %DB303.DBX6.0, 1 s
   "COMANDOS_MB-04-HS10" : Bool = PLC COMANDOS.MB-04-HS10 AT %DB303.DBX6.1, 1 s
   "COMANDOS_MB-04-HS11" : Bool = PLC COMANDOS.MB-04-HS11 AT %DB303.DBX6.2, 1 s
   "COMANDOS_MB-04-HS12" : Bool = PLC COMANDOS.MB-04-HS12 AT %DB303.DBX6.3, 1 s
   "COMANDOS_MB-04-HS13" : Bool = PLC COMANDOS.MB-04-HS13 AT %DB303.DBX6.4, 1 s
   "COMANDOS_MB-04-HS14" : Bool = PLC COMANDOS.MB-04-HS14 AT %DB303.DBX6.5, 1 s
   "COMANDOS_MB-04-HS15" : Bool = PLC COMANDOS.MB-04-HS15 AT %DB303.DBX6.6, 1 s
   "COMANDOS_MB-04-HS16" : Bool = PLC COMANDOS.MB-04-HS16 AT %DB303.DBX6.7, 1 s
   "COMANDOS_MB-04-HS1" : Bool = PLC COMANDOS.MB-04-HS1 AT %DB303.DBX7.0, 1 s
   "COMANDOS_MB-04-HS2" : Bool = PLC COMANDOS.MB-04-HS2 AT %DB303.DBX7.1, 1 s
   "COMANDOS_MB-04-HS3" : Bool = PLC COMANDOS.MB-04-HS3 AT %DB303.DBX7.2, 1 s
   "COMANDOS_MB-04-HS4" : Bool = PLC COMANDOS.MB-04-HS4 AT %DB303.DBX7.3, 1 s
   "COMANDOS_MB-04-HS5" : Bool = PLC COMANDOS.MB-04-HS5 AT %DB303.DBX7.4, 1 s
   "COMANDOS_MB-04-HS6" : Bool = PLC COMANDOS.MB-04-HS6 AT %DB303.DBX7.5, 1 s
   "COMANDOS_MB-04-HS7" : Bool = PLC COMANDOS.MB-04-HS7 AT %DB303.DBX7.6, 1 s
   "COMANDOS_MB-04-HS8" : Bool = PLC COMANDOS.MB-04-HS8 AT %DB303.DBX7.7, 1 s
   "COMANDOS_LIT_001-HS9" : Bool = PLC COMANDOS.LIT_001-HS9 AT %DB303.DBX8.0, 1 s
   "COMANDOS_LIT_001-HS10" : Bool = PLC COMANDOS.LIT_001-HS10 AT %DB303.DBX8.1, 1 s
   "COMANDOS_LIT_001-HS11" : Bool = PLC COMANDOS.LIT_001-HS11 AT %DB303.DBX8.2, 1 s
   "COMANDOS_LIT_001-HS12" : Bool = PLC COMANDOS.LIT_001-HS12 AT %DB303.DBX8.3, 1 s
   "COMANDOS_LIT_001-HS13" : Bool = PLC COMANDOS.LIT_001-HS13 AT %DB303.DBX8.4, 1 s
   "COMANDOS_LIT_001-HS14" : Bool = PLC COMANDOS.LIT_001-HS14 AT %DB303.DBX8.5, 1 s
   "COMANDOS_LIT_001-HS15" : Bool = PLC COMANDOS.LIT_001-HS15 AT %DB303.DBX8.6, 1 s
   "COMANDOS_LIT_001-HS16" : Bool = PLC COMANDOS.LIT_001-HS16 AT %DB303.DBX8.7, 1 s
   "COMANDOS_LIT_001-HSHH" : Bool = PLC COMANDOS.LIT_001-HSHH AT %DB303.DBX9.0, 1 s
   "COMANDOS_LIT_001-HSH" : Bool = PLC COMANDOS.LIT_001-HSH AT %DB303.DBX9.1, 1 s
   "COMANDOS_LIT_001-HSL" : Bool = PLC COMANDOS.LIT_001-HSL AT %DB303.DBX9.2, 1 s
   "COMANDOS_LIT_001-HSLL" : Bool = PLC COMANDOS.LIT_001-HSLL AT %DB303.DBX9.3, 1 s
   "COMANDOS_LIT_001-HSM" : Bool = PLC COMANDOS.LIT_001-HSM AT %DB303.DBX9.4, 1 s
   "COMANDOS_LIT_001-HS6" : Bool = PLC COMANDOS.LIT_001-HS6 AT %DB303.DBX9.5, 1 s
   "COMANDOS_LIT_001-HS7" : Bool = PLC COMANDOS.LIT_001-HS7 AT %DB303.DBX9.6, 1 s
   "COMANDOS_LIT_001-HS8" : Bool = PLC COMANDOS.LIT_001-HS8 AT %DB303.DBX9.7, 1 s
   "COMANDOS_PID-EEEB-HD" : Bool = PLC COMANDOS.PID-EEEB-HD AT %DB303.DBX10.1, 1 s
   "COMANDOS_PID-EEEB-HP" : Bool = PLC COMANDOS.PID-EEEB-HP AT %DB303.DBX10.2, 1 s
   "COMANDOS_PID-EEEB-HI" : Bool = PLC COMANDOS.PID-EEEB-HI AT %DB303.DBX10.3, 1 s
   "COMANDOS_PID-EEEB-HM" : Bool = PLC COMANDOS.PID-EEEB-HM AT %DB303.DBX12.2, 1 s

